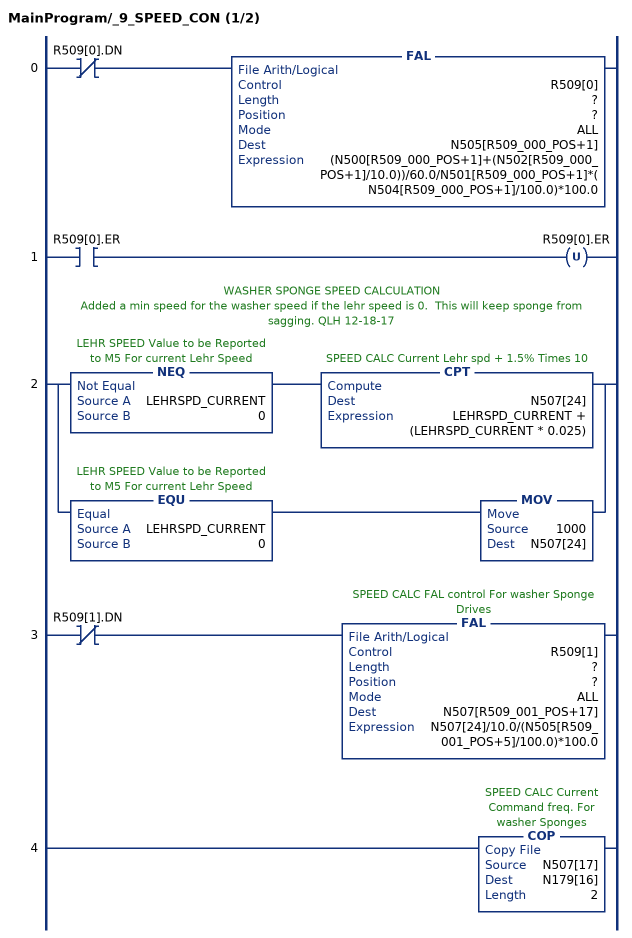
   0: XIO(R509[0].DN)FAL(R509[0],?,?,ALL,N505[R509_000_POS+1],(N500[R509_000_POS+1]+(N502[R509_000_POS+1]/10.0))/60.0/N501[R509_000_POS+1]*(N504[R509_000_POS+1]/100.0)*100.0);
   1: XIC(R509[0].ER)OTU(R509[0].ER);
   // WASHER SPONGE SPEED CALCULATION
   // Added a min speed for the washer speed if the lehr speed is 0.  This will keep sponge from sagging. QLH 12-18-17
   2: [NEQ(LEHRSPD_CURRENT,0) CPT(N507[24],LEHRSPD_CURRENT + (LEHRSPD_CURRENT * 0.025)) ,EQU(LEHRSPD_CURRENT,0) MOV(1000,N507[24]) ];
   3: XIO(R509[1].DN)FAL(R509[1],?,?,ALL,N507[R509_001_POS+17],N507[24]/10.0/(N505[R509_001_POS+5]/100.0)*100.0);
   4: COP(N507[17],N179[16],2);
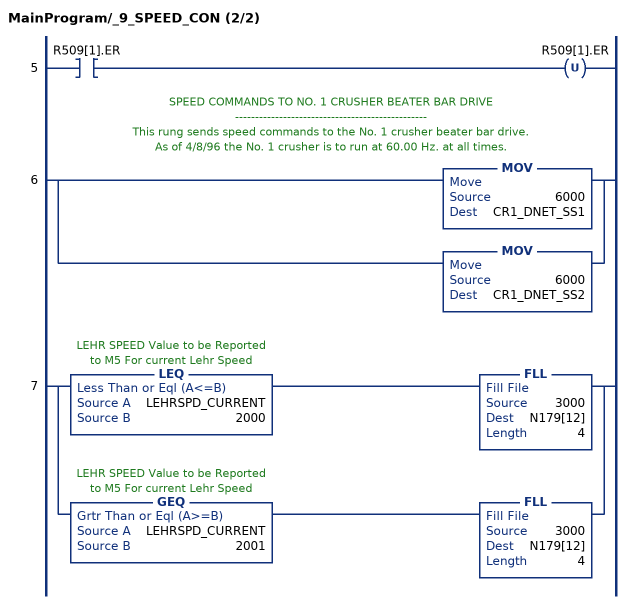
   5: XIC(R509[1].ER)OTU(R509[1].ER);
   // SPEED COMMANDS TO NO. 1 CRUSHER BEATER BAR DRIVE
   // ------------------------------------------------
   // This rung sends speed commands to the No. 1 crusher beater bar drive.
   // As of 4/8/96 the No. 1 crusher is to run at 60.00 Hz. at all times.
   6: [MOV(6000,CR1_DNET_SS1) ,MOV(6000,CR1_DNET_SS2) ];
   7: [LEQ(LEHRSPD_CURRENT,2000) FLL(3000,N179[12],4) ,GEQ(LEHRSPD_CURRENT,2001) FLL(3000,N179[12],4) ];
END_ROUTINE

ROUTINE _W_2_LADDER   (* ladder *)
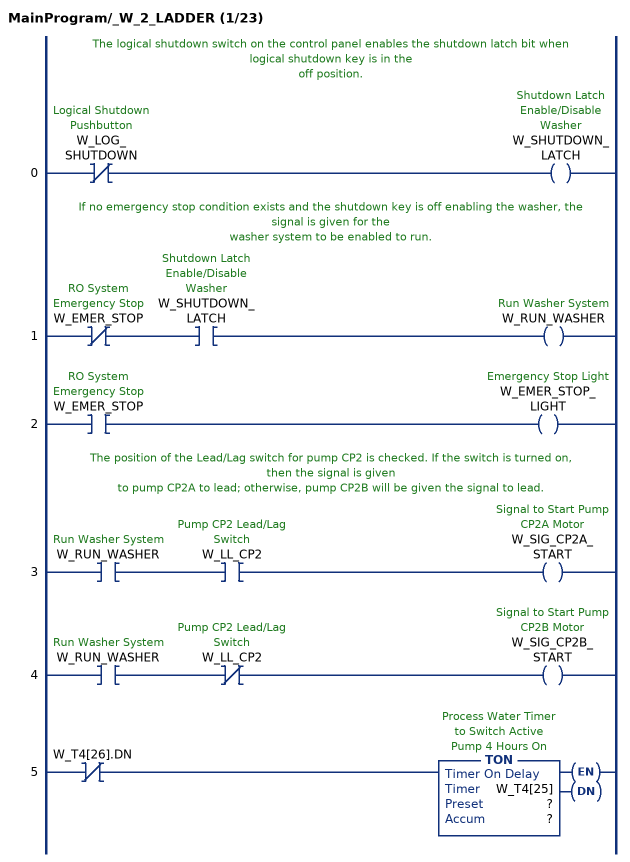
   // The logical shutdown switch on the control panel enables the shutdown latch bit when logical shutdown key is in the
   // off position.
   0: XIO(W_LOG_SHUTDOWN)OTE(W_SHUTDOWN_LATCH);
   // If no emergency stop condition exists and the shutdown key is off enabling the washer, the signal is given for the
   // washer system to be enabled to run.
   1: XIO(W_EMER_STOP)XIC(W_SHUTDOWN_LATCH)OTE(W_RUN_WASHER);
   2: XIC(W_EMER_STOP)OTE(W_EMER_STOP_LIGHT);
   // The position of the Lead/Lag switch for pump CP2 is checked. If the switch is turned on, then the signal is given
   // to pump CP2A to lead; otherwise, pump CP2B will be given the signal to lead.
   3: XIC(W_RUN_WASHER)XIC(W_LL_CP2)OTE(W_SIG_CP2A_START);
   4: XIC(W_RUN_WASHER)XIO(W_LL_CP2)OTE(W_SIG_CP2B_START);
   5: XIO(W_T4[26].DN)TON(W_T4[25],?,?);
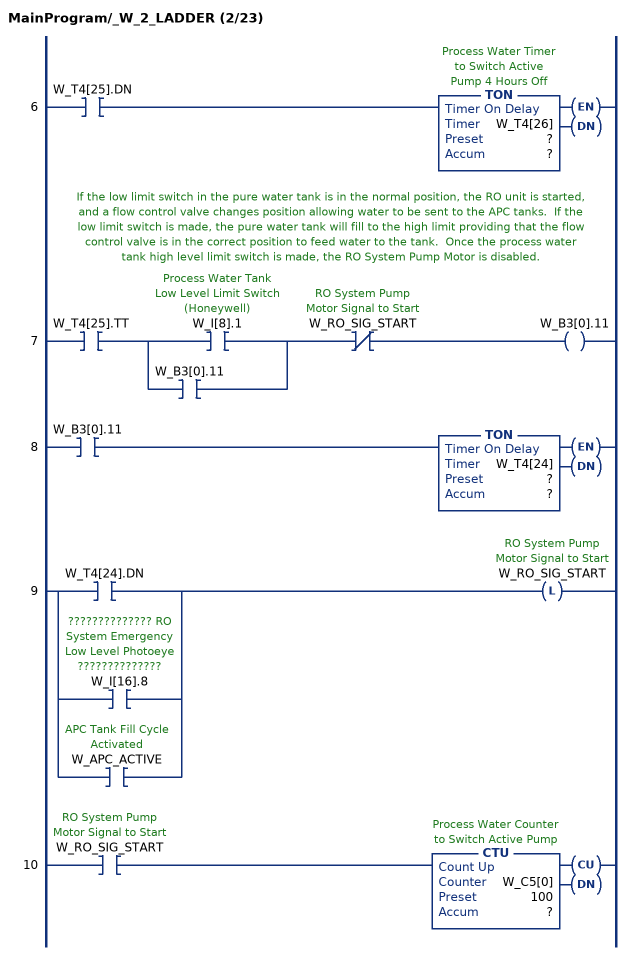
   6: XIC(W_T4[25].DN)TON(W_T4[26],?,?);
   // If the low limit switch in the pure water tank is in the normal position, the RO unit is started, and a flow control valve changes position allowing water to be sent to the APC tanks.  If the low limit switch is made, the pure water tank will fill to the high limit providing that the flow control valve is in the correct position to feed water to the tank.  Once the process water tank high level limit switch is made, the RO System Pump Motor is disabled.
   7: XIC(W_T4[25].TT)[XIC(W_I[8].1) ,XIC(W_B3[0].11) ]XIO(W_RO_SIG_START)OTE(W_B3[0].11);
   8: XIC(W_B3[0].11)TON(W_T4[24],?,?);
   9: [XIC(W_T4[24].DN) ,XIC(W_I[16].8) ,XIC(W_APC_ACTIVE) ]OTL(W_RO_SIG_START);
   10: XIC(W_RO_SIG_START)CTU(W_C5[0],?,?);
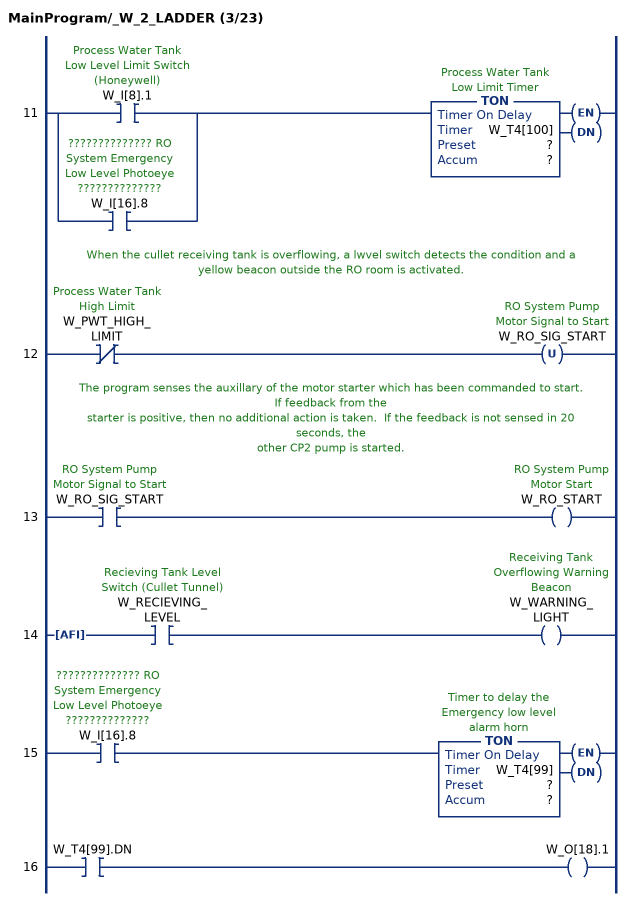
   11: [XIC(W_I[8].1) ,XIC(W_I[16].8) ]TON(W_T4[100],?,?);
   // When the cullet receiving tank is overflowing, a lwvel switch detects the condition and a yellow beacon outside the RO room is activated.
   12: XIO(W_PWT_HIGH_LIMIT)OTU(W_RO_SIG_START);
   // The program senses the auxillary of the motor starter which has been commanded to start.  If feedback from the
   // starter is positive, then no additional action is taken.  If the feedback is not sensed in 20 seconds, the
   // other CP2 pump is started.
   13: XIC(W_RO_SIG_START)OTE(W_RO_START);
   14: AFI()XIC(W_RECIEVING_LEVEL)OTE(W_WARNING_LIGHT);
   15: XIC(W_I[16].8)TON(W_T4[99],?,?);
   16: XIC(W_T4[99].DN)OTE(W_O[18].1);
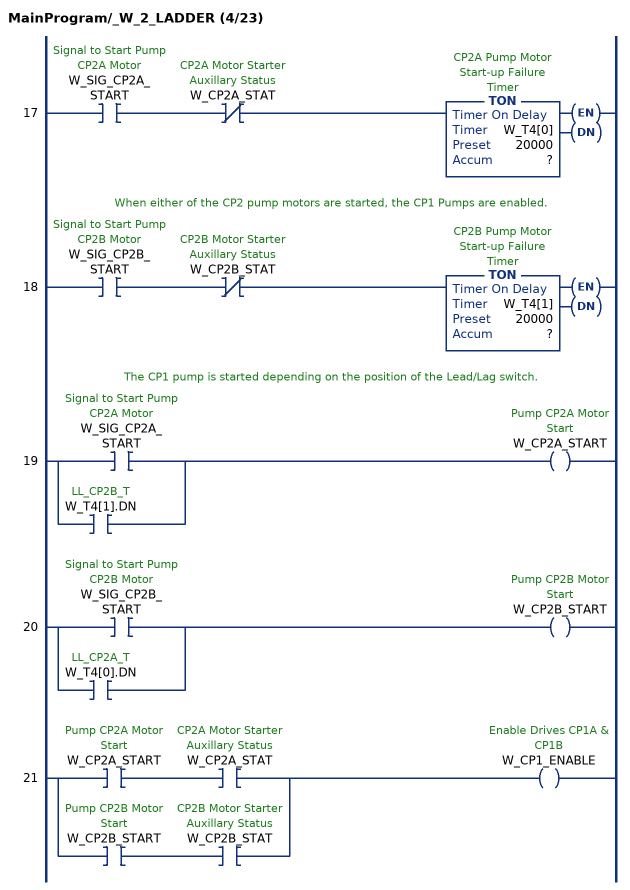
   17: XIC(W_SIG_CP2A_START)XIO(W_CP2A_STAT)TON(W_T4[0],?,?);
   // When either of the CP2 pump motors are started, the CP1 Pumps are enabled.
   18: XIC(W_SIG_CP2B_START)XIO(W_CP2B_STAT)TON(W_T4[1],?,?);
   // The CP1 pump is started depending on the position of the Lead/Lag switch.
   19: [XIC(W_SIG_CP2A_START) ,XIC(W_T4[1].DN) ]OTE(W_CP2A_START);
   20: [XIC(W_SIG_CP2B_START) ,XIC(W_T4[0].DN) ]OTE(W_CP2B_START);
   21: [XIC(W_CP2A_START) XIC(W_CP2A_STAT) ,XIC(W_CP2B_START) XIC(W_CP2B_STAT) ]OTE(W_CP1_ENABLE);
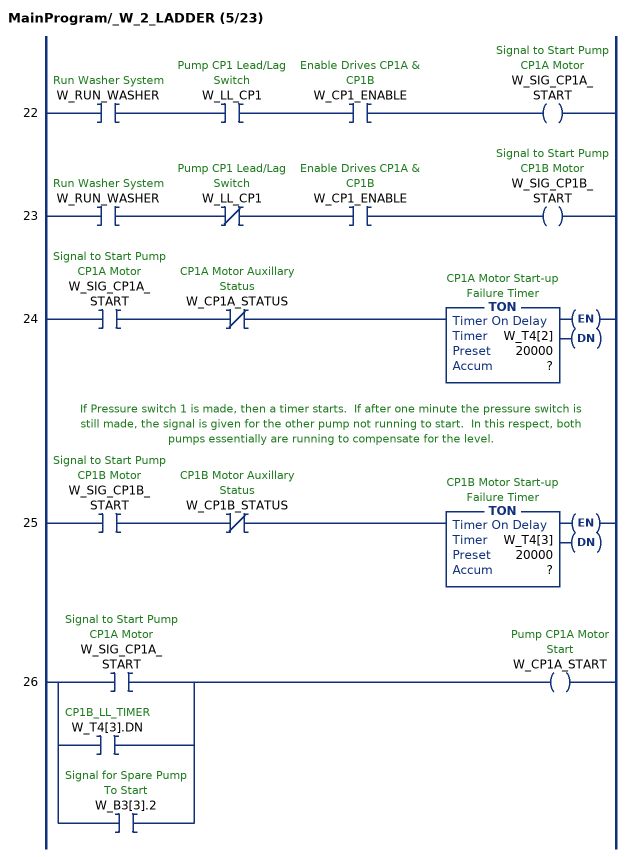
   22: XIC(W_RUN_WASHER)XIC(W_LL_CP1)XIC(W_CP1_ENABLE)OTE(W_SIG_CP1A_START);
   23: XIC(W_RUN_WASHER)XIO(W_LL_CP1)XIC(W_CP1_ENABLE)OTE(W_SIG_CP1B_START);
   24: XIC(W_SIG_CP1A_START)XIO(W_CP1A_STATUS)TON(W_T4[2],?,?);
   // If Pressure switch 1 is made, then a timer starts.  If after one minute the pressure switch is still made, the signal is given for the other pump not running to start.  In this respect, both pumps essentially are running to compensate for the level.
   25: XIC(W_SIG_CP1B_START)XIO(W_CP1B_STATUS)TON(W_T4[3],?,?);
   26: [XIC(W_SIG_CP1A_START) ,XIC(W_T4[3].DN) ,XIC(W_B3[3].2) ]OTE(W_CP1A_START);
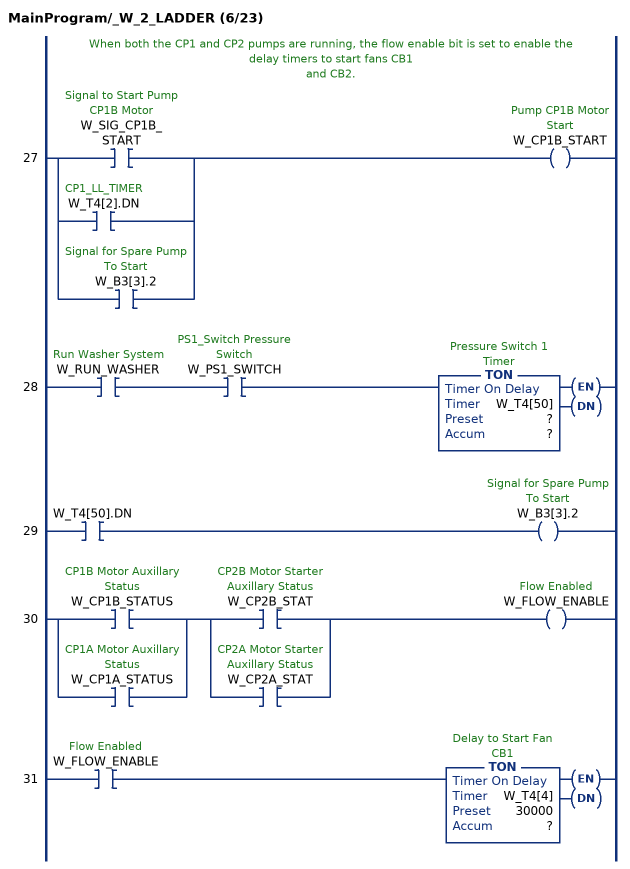
   // When both the CP1 and CP2 pumps are running, the flow enable bit is set to enable the delay timers to start fans CB1
   // and CB2.
   27: [XIC(W_SIG_CP1B_START) ,XIC(W_T4[2].DN) ,XIC(W_B3[3].2) ]OTE(W_CP1B_START);
   28: XIC(W_RUN_WASHER)XIC(W_PS1_SWITCH)TON(W_T4[50],?,?);
   29: XIC(W_T4[50].DN)OTE(W_B3[3].2);
   30: [XIC(W_CP1B_STATUS) ,XIC(W_CP1A_STATUS) ][XIC(W_CP2B_STAT) ,XIC(W_CP2A_STAT) ]OTE(W_FLOW_ENABLE);
   31: XIC(W_FLOW_ENABLE)TON(W_T4[4],?,?);
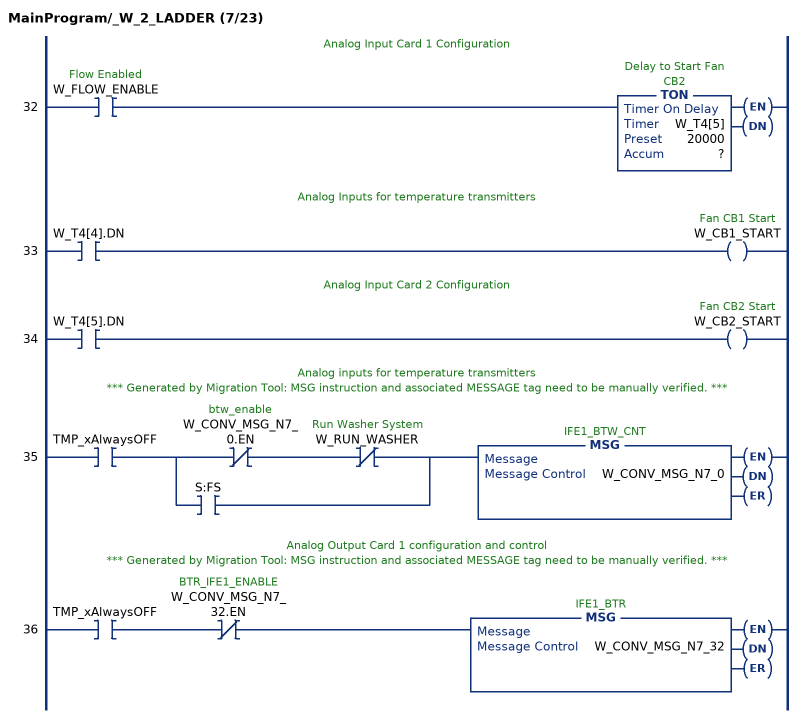
   // Analog Input Card 1 Configuration
   32: XIC(W_FLOW_ENABLE)TON(W_T4[5],?,?);
   // Analog Inputs for temperature transmitters
   33: XIC(W_T4[4].DN)OTE(W_CB1_START);
   // Analog Input Card 2 Configuration
   34: XIC(W_T4[5].DN)OTE(W_CB2_START);
   // Analog inputs for temperature transmitters
   // *** Generated by Migration Tool: MSG instruction and associated MESSAGE tag need to be manually verified. ***
   35: XIC(TMP_xAlwaysOFF)[XIO(W_CONV_MSG_N7_0.EN) XIO(W_RUN_WASHER) ,XIC(S:FS) ]MSG(W_CONV_MSG_N7_0);
   // Analog Output Card 1 configuration and control
   // *** Generated by Migration Tool: MSG instruction and associated MESSAGE tag need to be manually verified. ***
   36: XIC(TMP_xAlwaysOFF)XIO(W_CONV_MSG_N7_32.EN)MSG(W_CONV_MSG_N7_32);
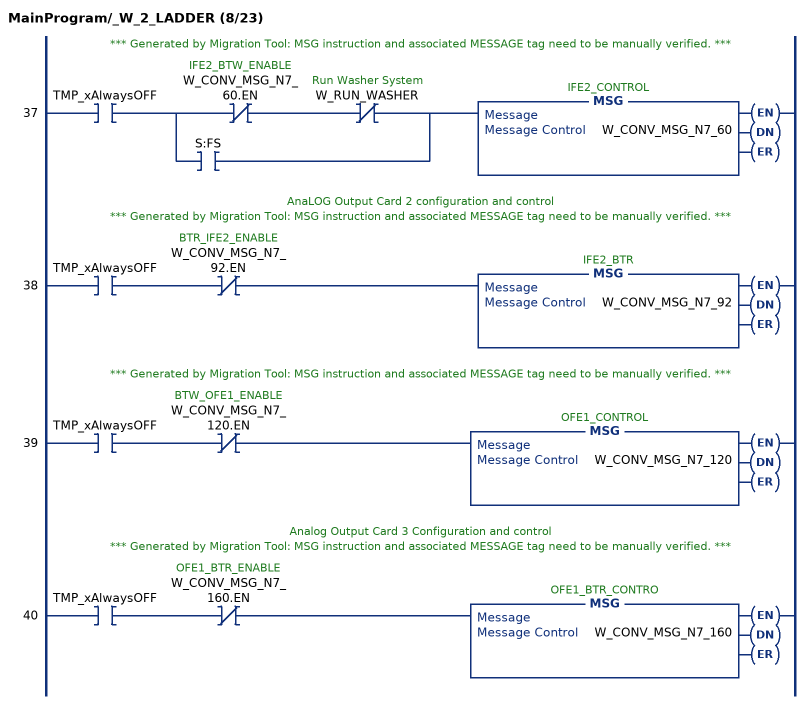
   // *** Generated by Migration Tool: MSG instruction and associated MESSAGE tag need to be manually verified. ***
   37: XIC(TMP_xAlwaysOFF)[XIO(W_CONV_MSG_N7_60.EN) XIO(W_RUN_WASHER) ,XIC(S:FS) ]MSG(W_CONV_MSG_N7_60);
   // AnaLOG Output Card 2 configuration and control
   // *** Generated by Migration Tool: MSG instruction and associated MESSAGE tag need to be manually verified. ***
   38: XIC(TMP_xAlwaysOFF)XIO(W_CONV_MSG_N7_92.EN)MSG(W_CONV_MSG_N7_92);
   // *** Generated by Migration Tool: MSG instruction and associated MESSAGE tag need to be manually verified. ***
   39: XIC(TMP_xAlwaysOFF)XIO(W_CONV_MSG_N7_120.EN)MSG(W_CONV_MSG_N7_120);
   // Analog Output Card 3 Configuration and control
   // *** Generated by Migration Tool: MSG instruction and associated MESSAGE tag need to be manually verified. ***
   40: XIC(TMP_xAlwaysOFF)XIO(W_CONV_MSG_N7_160.EN)MSG(W_CONV_MSG_N7_160);
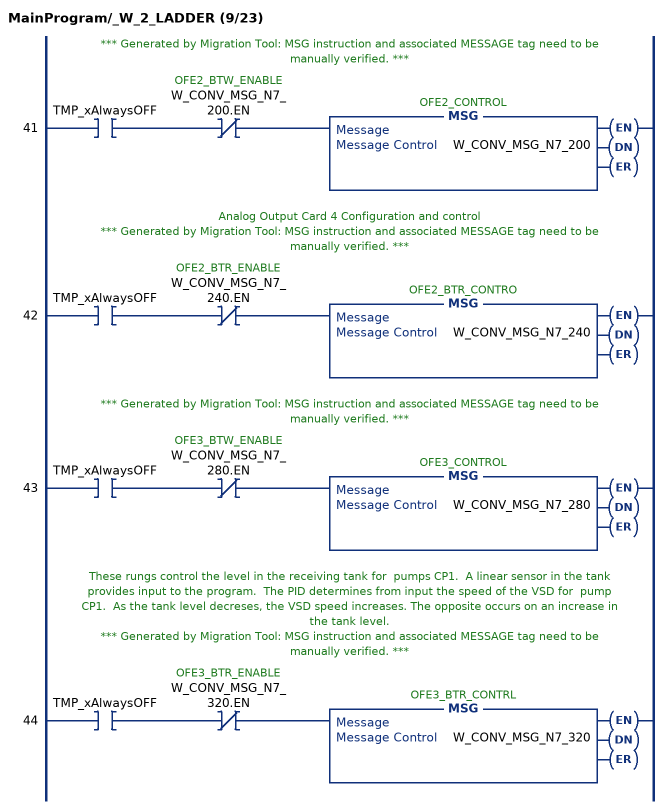
   // *** Generated by Migration Tool: MSG instruction and associated MESSAGE tag need to be manually verified. ***
   41: XIC(TMP_xAlwaysOFF)XIO(W_CONV_MSG_N7_200.EN)MSG(W_CONV_MSG_N7_200);
   // Analog Output Card 4 Configuration and control
   // *** Generated by Migration Tool: MSG instruction and associated MESSAGE tag need to be manually verified. ***
   42: XIC(TMP_xAlwaysOFF)XIO(W_CONV_MSG_N7_240.EN)MSG(W_CONV_MSG_N7_240);
   // *** Generated by Migration Tool: MSG instruction and associated MESSAGE tag need to be manually verified. ***
   43: XIC(TMP_xAlwaysOFF)XIO(W_CONV_MSG_N7_280.EN)MSG(W_CONV_MSG_N7_280);
   // These rungs control the level in the receiving tank for  pumps CP1.  A linear sensor in the tank provides input to the program.  The PID determines from input the speed of the VSD for  pump CP1.  As the tank level decreses, the VSD speed increases. The opposite occurs on an increase in the tank level.
   // *** Generated by Migration Tool: MSG instruction and associated MESSAGE tag need to be manually verified. ***
   44: XIC(TMP_xAlwaysOFF)XIO(W_CONV_MSG_N7_320.EN)MSG(W_CONV_MSG_N7_320);
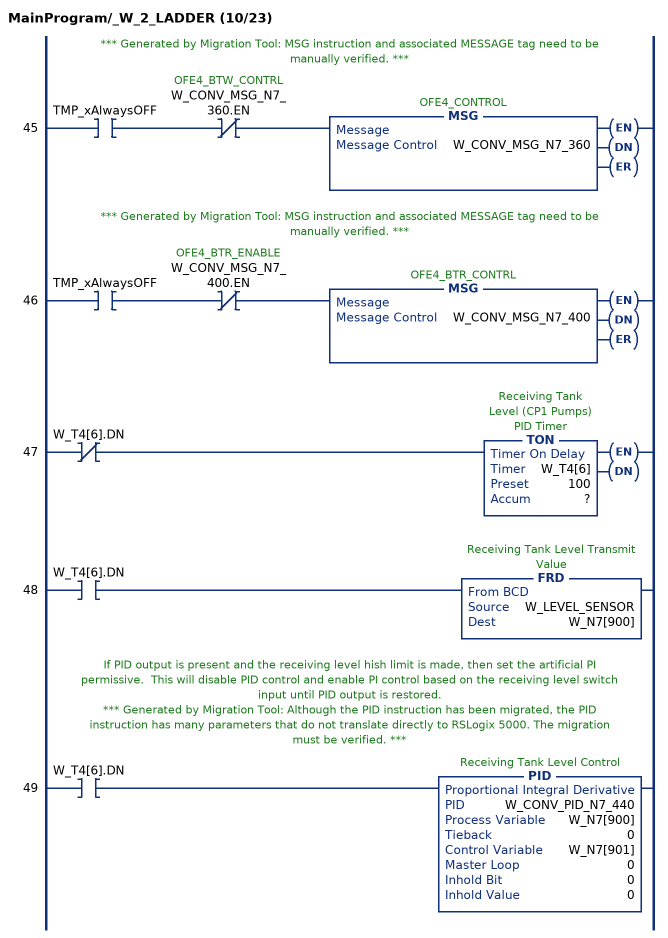
   // *** Generated by Migration Tool: MSG instruction and associated MESSAGE tag need to be manually verified. ***
   45: XIC(TMP_xAlwaysOFF)XIO(W_CONV_MSG_N7_360.EN)MSG(W_CONV_MSG_N7_360);
   // *** Generated by Migration Tool: MSG instruction and associated MESSAGE tag need to be manually verified. ***
   46: XIC(TMP_xAlwaysOFF)XIO(W_CONV_MSG_N7_400.EN)MSG(W_CONV_MSG_N7_400);
   47: XIO(W_T4[6].DN)TON(W_T4[6],?,?);
   48: XIC(W_T4[6].DN)FRD(W_LEVEL_SENSOR,W_N7[900]);
   // If PID output is present and the receiving level hish limit is made, then set the artificial PI permissive.  This will disable PID control and enable PI control based on the receiving level switch input until PID output is restored.
   // *** Generated by Migration Tool: Although the PID instruction has been migrated, the PID instruction has many parameters that do not translate directly to RSLogix 5000. The migration must be verified. ***
   49: XIC(W_T4[6].DN)PID(W_CONV_PID_N7_440,W_N7[900],0,W_N7[901],0,0,0);
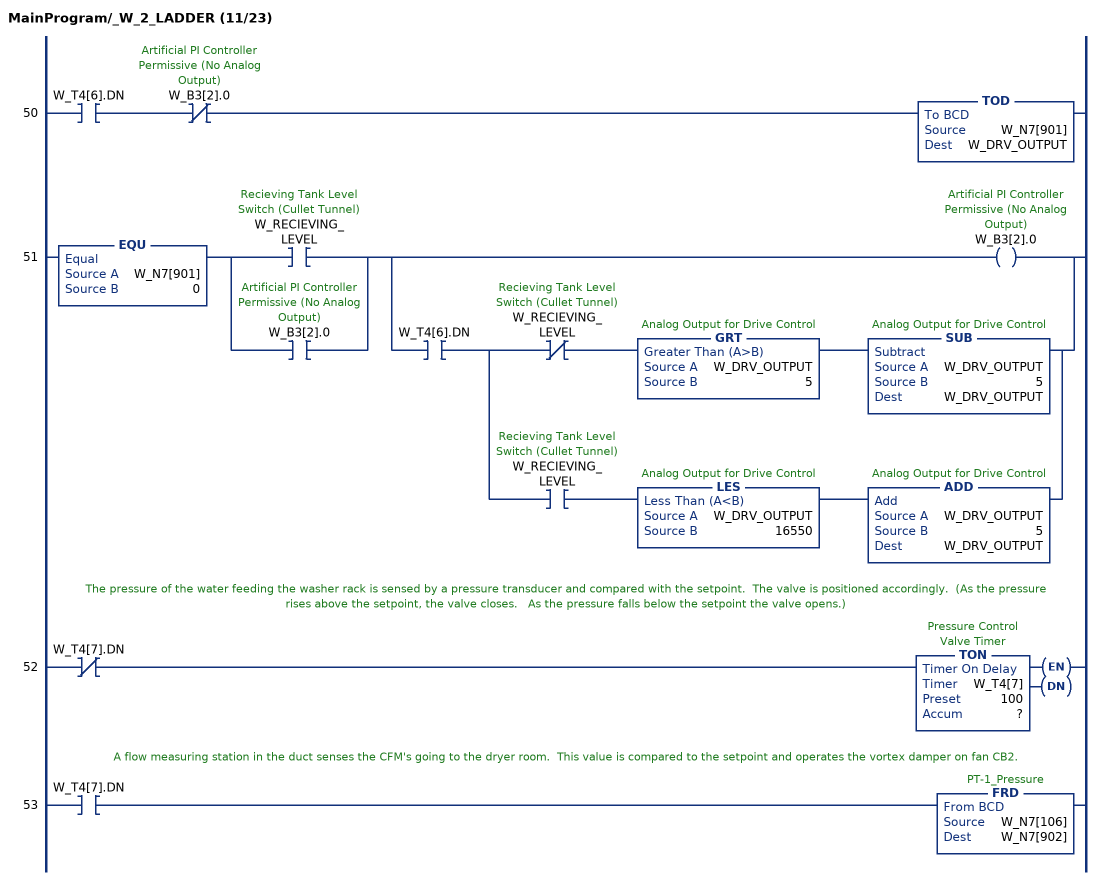
   50: XIC(W_T4[6].DN)XIO(W_B3[2].0)TOD(W_N7[901],W_DRV_OUTPUT);
   51: EQU(W_N7[901],0)[XIC(W_RECIEVING_LEVEL) ,XIC(W_B3[2].0) ][OTE(W_B3[2].0) ,XIC(W_T4[6].DN) [XIO(W_RECIEVING_LEVEL) GRT(W_DRV_OUTPUT,5) SUB(W_DRV_OUTPUT,5,W_DRV_OUTPUT) ,XIC(W_RECIEVING_LEVEL) LES(W_DRV_OUTPUT,16550) ADD(W_DRV_OUTPUT,5,W_DRV_OUTPUT) ] ];
   // The pressure of the water feeding the washer rack is sensed by a pressure transducer and compared with the setpoint.  The valve is positioned accordingly.  (As the pressure rises above the setpoint, the valve closes.   As the pressure falls below the setpoint the valve opens.)
   52: XIO(W_T4[7].DN)TON(W_T4[7],?,?);
   // A flow measuring station in the duct senses the CFM's going to the dryer room.  This value is compared to the setpoint and operates the vortex damper on fan CB2.
   53: XIC(W_T4[7].DN)FRD(W_N7[106],W_N7[902]);
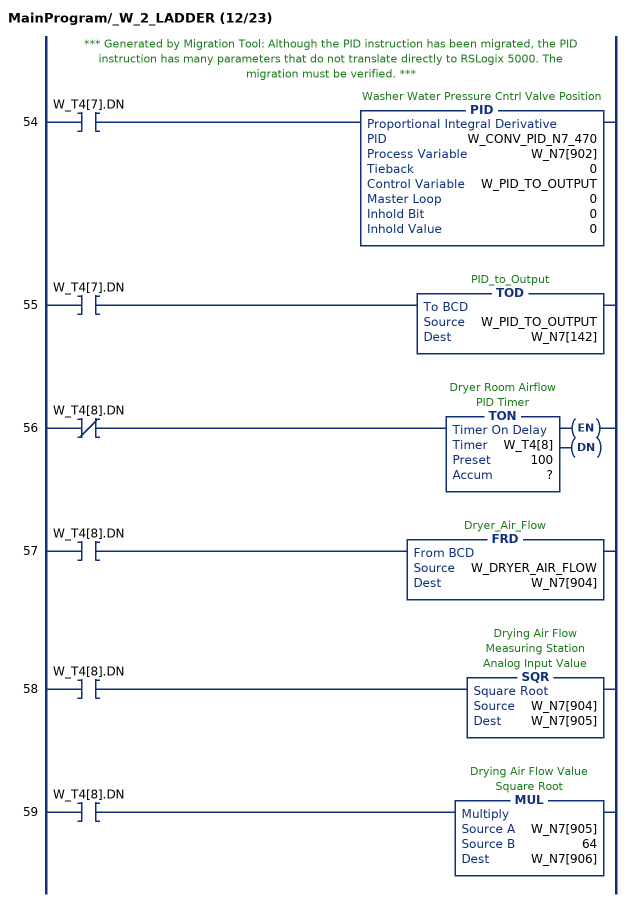
   // *** Generated by Migration Tool: Although the PID instruction has been migrated, the PID instruction has many parameters that do not translate directly to RSLogix 5000. The migration must be verified. ***
   54: XIC(W_T4[7].DN)PID(W_CONV_PID_N7_470,W_N7[902],0,W_PID_TO_OUTPUT,0,0,0);
   55: XIC(W_T4[7].DN)TOD(W_PID_TO_OUTPUT,W_N7[142]);
   56: XIO(W_T4[8].DN)TON(W_T4[8],?,?);
   57: XIC(W_T4[8].DN)FRD(W_DRYER_AIR_FLOW,W_N7[904]);
   58: XIC(W_T4[8].DN)SQR(W_N7[904],W_N7[905]);
   59: XIC(W_T4[8].DN)MUL(W_N7[905],64,W_N7[906]);
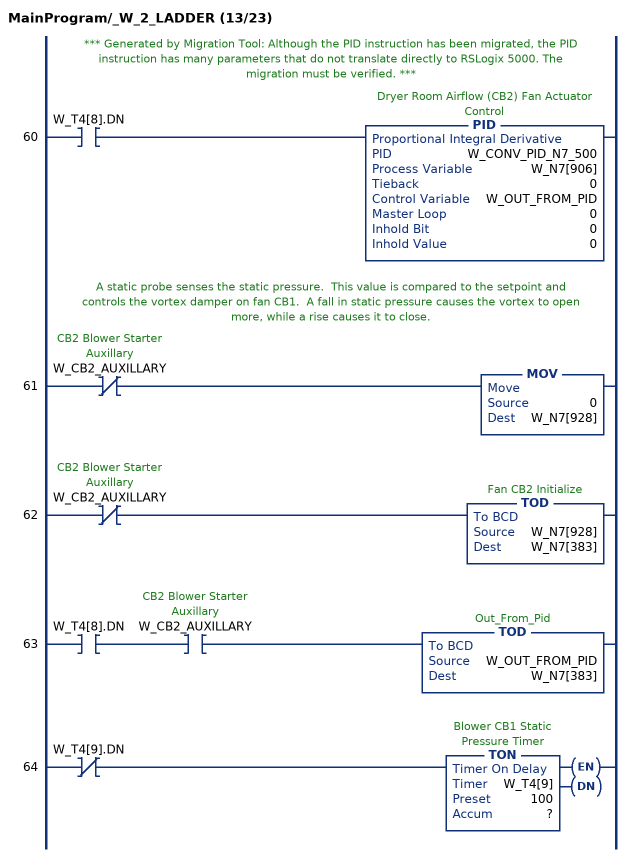
   // *** Generated by Migration Tool: Although the PID instruction has been migrated, the PID instruction has many parameters that do not translate directly to RSLogix 5000. The migration must be verified. ***
   60: XIC(W_T4[8].DN)PID(W_CONV_PID_N7_500,W_N7[906],0,W_OUT_FROM_PID,0,0,0);
   // A static probe senses the static pressure.  This value is compared to the setpoint and controls the vortex damper on fan CB1.  A fall in static pressure causes the vortex to open more, while a rise causes it to close.
   61: XIO(W_CB2_AUXILLARY)MOV(0,W_N7[928]);
   62: XIO(W_CB2_AUXILLARY)TOD(W_N7[928],W_N7[383]);
   63: XIC(W_T4[8].DN)XIC(W_CB2_AUXILLARY)TOD(W_OUT_FROM_PID,W_N7[383]);
   64: XIO(W_T4[9].DN)TON(W_T4[9],?,?);
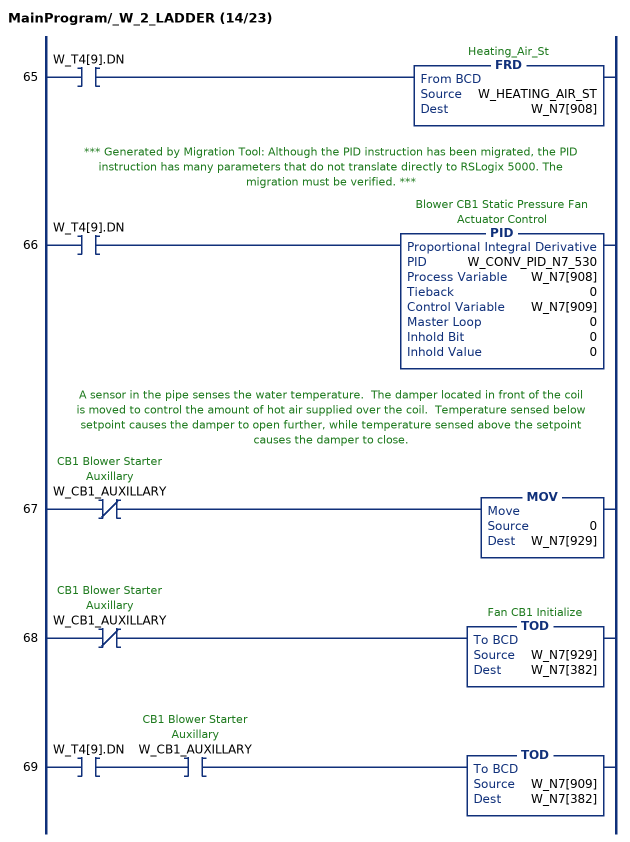
   65: XIC(W_T4[9].DN)FRD(W_HEATING_AIR_ST,W_N7[908]);
   // *** Generated by Migration Tool: Although the PID instruction has been migrated, the PID instruction has many parameters that do not translate directly to RSLogix 5000. The migration must be verified. ***
   66: XIC(W_T4[9].DN)PID(W_CONV_PID_N7_530,W_N7[908],0,W_N7[909],0,0,0);
   // A sensor in the pipe senses the water temperature.  The damper located in front of the coil is moved to control the amount of hot air supplied over the coil.  Temperature sensed below setpoint causes the damper to open further, while temperature sensed above the setpoint causes the damper to close.
   67: XIO(W_CB1_AUXILLARY)MOV(0,W_N7[929]);
   68: XIO(W_CB1_AUXILLARY)TOD(W_N7[929],W_N7[382]);
   69: XIC(W_T4[9].DN)XIC(W_CB1_AUXILLARY)TOD(W_N7[909],W_N7[382]);
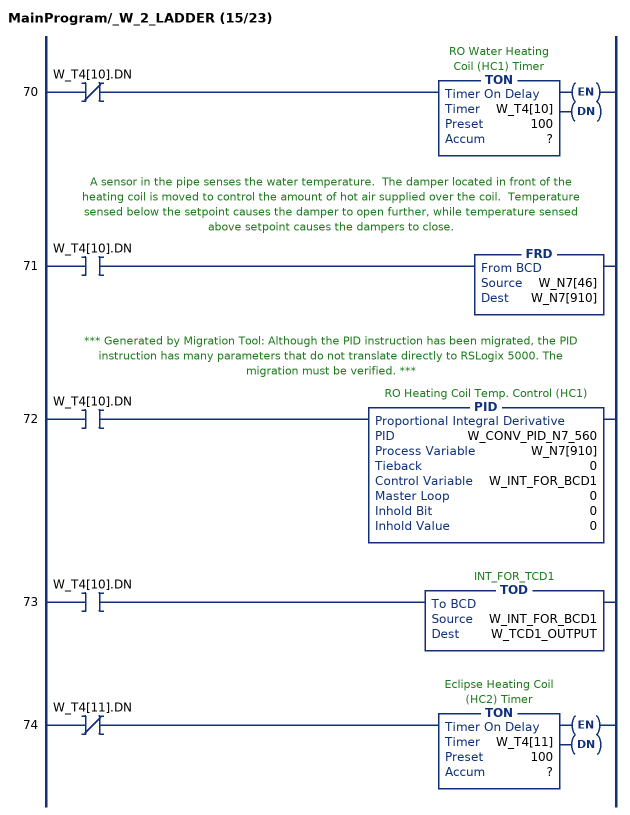
   70: XIO(W_T4[10].DN)TON(W_T4[10],?,?);
   // A sensor in the pipe senses the water temperature.  The damper located in front of the heating coil is moved to control the amount of hot air supplied over the coil.  Temperature sensed below the setpoint causes the damper to open further, while temperature sensed above setpoint causes the dampers to close.
   71: XIC(W_T4[10].DN)FRD(W_N7[46],W_N7[910]);
   // *** Generated by Migration Tool: Although the PID instruction has been migrated, the PID instruction has many parameters that do not translate directly to RSLogix 5000. The migration must be verified. ***
   72: XIC(W_T4[10].DN)PID(W_CONV_PID_N7_560,W_N7[910],0,W_INT_FOR_BCD1,0,0,0);
   73: XIC(W_T4[10].DN)TOD(W_INT_FOR_BCD1,W_TCD1_OUTPUT);
   74: XIO(W_T4[11].DN)TON(W_T4[11],?,?);
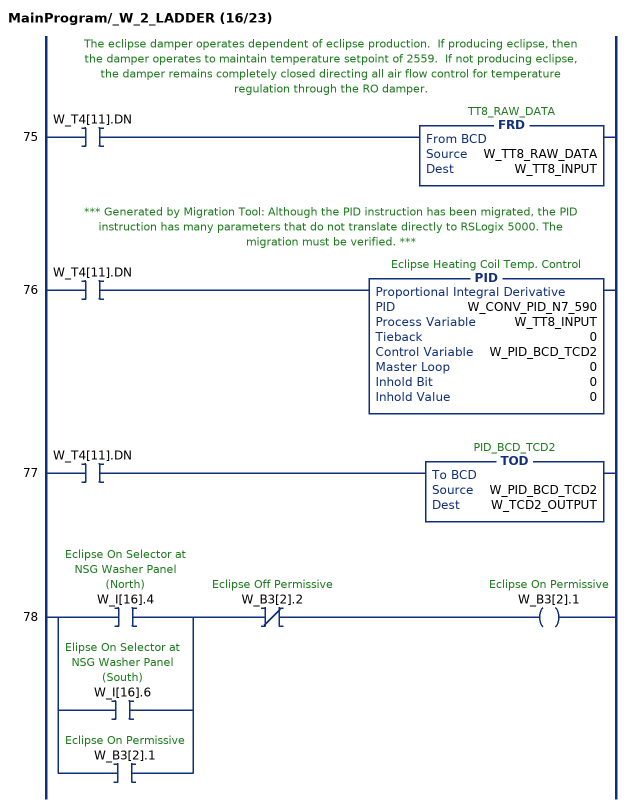
   // The eclipse damper operates dependent of eclipse production.  If producing eclipse, then the damper operates to maintain temperature setpoint of 2559.  If not producing eclipse, the damper remains completely closed directing all air flow control for temperature regulation through the RO damper.
   75: XIC(W_T4[11].DN)FRD(W_TT8_RAW_DATA,W_TT8_INPUT);
   // *** Generated by Migration Tool: Although the PID instruction has been migrated, the PID instruction has many parameters that do not translate directly to RSLogix 5000. The migration must be verified. ***
   76: XIC(W_T4[11].DN)PID(W_CONV_PID_N7_590,W_TT8_INPUT,0,W_PID_BCD_TCD2,0,0,0);
   77: XIC(W_T4[11].DN)TOD(W_PID_BCD_TCD2,W_TCD2_OUTPUT);
   78: [XIC(W_I[16].4) ,XIC(W_I[16].6) ,XIC(W_B3[2].1) ]XIO(W_B3[2].2)OTE(W_B3[2].1);
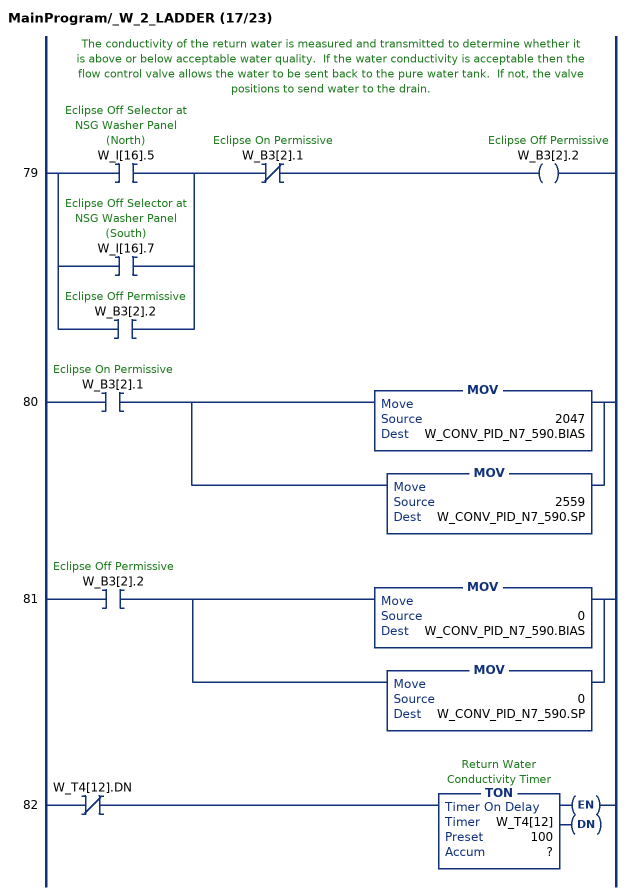
   // The conductivity of the return water is measured and transmitted to determine whether it is above or below acceptable water quality.  If the water conductivity is acceptable then the flow control valve allows the water to be sent back to the pure water tank.  If not, the valve positions to send water to the drain.
   79: [XIC(W_I[16].5) ,XIC(W_I[16].7) ,XIC(W_B3[2].2) ]XIO(W_B3[2].1)OTE(W_B3[2].2);
   80: XIC(W_B3[2].1)[MOV(2047,W_CONV_PID_N7_590.BIAS) ,MOV(2559,W_CONV_PID_N7_590.SP) ];
   81: XIC(W_B3[2].2)[MOV(0,W_CONV_PID_N7_590.BIAS) ,MOV(0,W_CONV_PID_N7_590.SP) ];
   82: XIO(W_T4[12].DN)TON(W_T4[12],?,?);
